// Mitsubishi GX Works2 project: ZhaoQing_FenRong_Debug   PLC: Q06UDEH

TYPE ShuttleCarIO : STRUCT
  xReady : BOOL;  (* 准备就绪 *)
  xForward : BOOL;  (* 正转 *)
  xBackward : BOOL;  (* 反转 *)
  iCurrentPos : INT;  (* 当前位置 *)
  iDestinationPos : INT;  (* 目标位置 *)
  xCW : BOOL;  (* 正转输出 *)
  xCCW : BOOL;  (* 反转输出 *)
  xBrake : BOOL;  (* 刹车 *)
  xHomeSwitch : BOOL;  (* 零位接近开关 *)
  xPosLimit : BOOL;  (* 正限位 *)
  xNegLimit : BOOL;  (* 负限位 *)
  xMDIExe : BOOL;  (* MDI开始 *)
  xMDIDone : BOOL;  (* MDI 完成 *)
  xPassLimit : BOOL;  (* 限位屏蔽 *)
  xPosLimitCatch : BOOL;  (* 正限位捕捉 *)
  xNegLimitCatch : BOOL;  (* 负限位捕捉 *)
  xHomeExe : BOOL;  (* 开始寻零 *)
  xHomeDone : BOOL;  (* 寻零完成 *)
  xHomeBusy : BOOL;  (* 寻零中 *)
  xHomeFailed : BOOL;  (* 寻零失败 *)
  xBusy : BOOL;  (* 工作中 *)
  tArriveDelay : TIME;  (* 到位延时 *)
  xCylinder : BOOL;  (* 气缸控制 *)
  tBrakeDelay : TIME;  (* 抱闸延时 *)
  xPauseRamp : BOOL;  (* 暂停减速斜坡标志位 *)
  xPresentDetect1 : BOOL;  (* 物料有无检测1 *)
  xPresentDetect2 : BOOL;  (* 物料有无检测2 *)
  xOvertimeAlarm : BOOL;  (* 超时报警 *)
  tSetOverTime : TIME;  (* 设置超时时间 *)
  xLooseDetect : BOOL;  (* 松绳检测 *)
  xLooseAlarm : BOOL;  (* 松绳报警 *)
END_STRUCT END_TYPE

TYPE SwitchIO : STRUCT
  xLiftCylinderRetractDetect : BOOL;
  xLiftCylinderExtendDetect : BOOL;
  xLiftCylinderRetract : BOOL;
  xLiftCylinderExtend : BOOL;
  xEntryBarCylinderRetract : BOOL;
  xLiftCylinderExtendInit : BOOL;
  xEntryEnable : BOOL;
  xExitEnable : BOOL;
  xExitBarCylinderRetract : BOOL;
  xSwithEnable : BOOL;
  xLiftCylinderRetractButton : BOOL;
  xLiftCylinderExtendButton : BOOL;
  xEntryBarCylinderRetractButton : BOOL;
  xExitBarCylinderRetractButton : BOOL;
END_STRUCT END_TYPE

TYPE BarCylinderIO : STRUCT
  xPresentSwitch : BOOL;  (* 行程开关 *)
  xBarCylinder : BOOL;  (* 阻挡气缸 *)
  xEmpty : BOOL;  (* 为空指示 *)
  xTransportMotorCW : BOOL;  (* 输送电机正转 *)
  xUnload : BOOL;  (* 下料 *)
  xBarCylinderButton : BOOL;  (* 阻挡气缸 *)
  xTransportMotorCWButton : BOOL;  (* 输送电机正转按钮 *)
  xLoad : BOOL;  (* 上料 *)
  xNextRun : BOOL;  (* 下位设备开始运行 *)
  xTransportMotorCCWButton : BOOL;  (* 输送电机反转按钮 *)
  xTransportMotorCCW : BOOL;  (* 输送电机反转 *)
  iProductCategory : INT;  (* 产品种类 *)
  tLoadDelay : TIME;  (* 上料延时 *)
END_STRUCT END_TYPE

TYPE ConveyorIO : STRUCT
  iProductCategory : INT;  (* 产品类型0：无料1：正极  2：负极 3：隔膜 4：空料架 *)
  xCWPresent : BOOL;  (* 正转检测有无传感器 *)
  xCCWPresent : BOOL;  (* 反转检测有无传感器 *)
  xLoad : BOOL;  (* 上料请求 *)
  xUnload : BOOL;  (* 下料请求 *)
  xMotorCW : BOOL;  (* 电机正转 *)
  xMotorCCW : BOOL;  (* 电机反转 *)
  xEmpty : BOOL;  (* 线体状态为空 *)
  xNextRun : BOOL;  (* 下段线体运行 *)
  xUnloadCCW : BOOL;  (* 下料为反转 *)
  xloadCCW : BOOL;  (* 上料为反转 *)
  xLeave : BOOL;  (* 已经离开 *)
  xForward : BOOL;  (* 正转手动 *)
  xBackward : BOOL;  (* 反转手动 *)
  xBusy : BOOL;  (* 工作中 *)
  tLoadDelay : TIME;  (* 进入延时设置 *)
  xPutInto : BOOL;  (* 线体直接投入物料 *)
  xUnloadAlarm : BOOL;  (* 下料报警 *)
  xPosLimit : BOOL;  (* 正限位 *)
  xNegLimit : BOOL;  (* 负限位 *)
  xOverWidthAlarm : BOOL;  (* 超宽报警 *)
  xLimitAlarrm : BOOL;  (* 限位报警 *)
  iDeviceID : INT;  (* 线体ID *)
  xSizeDeficientDetect : BOOL;  (* 尺寸不足检测标志位 *)
END_STRUCT END_TYPE

TYPE RGVCommunication : STRUCT
  xFullLoadRequest : BOOL;  (* 满框上料请求 *)
  xFullUnloadRequest : BOOL;  (* 满框下料请求 *)
  xEmptyLoadRequest : BOOL;  (* 空框上料请求 *)
  xEmptyUnloadRequest : BOOL;  (* 空框下料请求 *)
  xFullLoadRequestAkn : BOOL;  (* 满框上料请求确认 *)
  xFullUnloadRequestAkn : BOOL;  (* 满框下料请求确认 *)
  xEmptyLoadRequestAkn : BOOL;  (* 空框上料请求确认 *)
  xEmptyUnloadRequestAkn : BOOL;  (* 空框下料请求确认 *)
  xFullLoadComplete : BOOL;  (* 满框上料完成 *)
  xFullUnloadComplete : BOOL;  (* 满框下料完成 *)
  xEmptyLoadComplete : BOOL;  (* 空框上料完成 *)
  xEmptyUnloadComplete : BOOL;  (* 空框下料完成 *)
  xFullLoadCompleteAkn : BOOL;  (* 满框上料完成确认 *)
  xFullUnloadCompleteAkn : BOOL;  (* 满框下料完成确认 *)
  xEmptyLoadCompleteAkn : BOOL;  (* 空框上料完成确认 *)
  xEmptyUnloadCompleteAkn : BOOL;  (* 空框下料完成确认 *)
  xMdiExe : BOOL;  (* RGV 执行 *)
  xMdiDone : BOOL;  (* RGV 执行完成 *)
  iCurrentPostion : INT;  (* RGV当前位置 *)
  iDestinationPos : INT;  (* RGV目标位置 *)
  xEmpty1 : BOOL;
  xNextRun1 : BOOL;
  xEmpty2 : BOOL;
  xNextRun2 : BOOL;
  xLoad1 : BOOL;
  xUnload1 : BOOL;
  xLoad2 : BOOL;
  xUnload2 : BOOL;
  xCollisionAlarm : BOOL;  (* 干涉报警 *)
  xRemoteReset : BOOL;  (* 远程复位 *)
  xAuto : BOOL;  (* 自动 *)
END_STRUCT END_TYPE

TYPE Stub : STRUCT
  xLoadRequest : BOOL;
  xLoadRequestAkn : BOOL;
  xUnloadRequest : BOOL;
  xUnloadRequestAkn : BOOL;
END_STRUCT END_TYPE

// global labels: Global1
VAR_GLOBAL
  g_xAuto AT M11 : BOOL;
  g_xManual : BOOL;
  g_xEStop AT X33 : BOOL;
  g_xReset AT X30 : BOOL;
  g_xStackLampRed AT Y230 : BOOL;
  g_xStackLampAmber AT Y231 : BOOL;
  g_xStackLampGreen AT Y232 : BOOL;
  g_xBuzzer AT Y233 : BOOL;
  g_xStop AT M2 : BOOL;
  g_xLocalAutoStart AT M1 : BOOL;
  g_xRemoteAutoStart AT M0 : BOOL;
  g_xRemoteAuto AT M10 : BOOL;
  g_iState AT D40 : INT;
  g_iLocalAutoStep : INT;
  g_xImport1Force AT M141 : BOOL;  (* 常温库1巷道单框强制入库 *)
  g_xImport2Force AT M142 : BOOL;  (* 常温库2巷道单框强制入库 *)
  g_xImport3Force AT M143 : BOOL;  (* 常温库3巷道单框强制入库 *)
  g_xForbidLifter7 AT M146 : BOOL;  (* 禁用提升机7 *)
  g_xResetSingle AT M4 : BOOL;  (* 单线体复位 *)
  g_iDeviceIDSelect AT D0 : INT;
  g_xPause AT M3 : BOOL;  (* 暂停 *)
  g_xAlarm : BOOL;  (* 报警 *)
  g_xCommissioning : BOOL;  (* 调试模式 *)
END_VAR

// global labels: Global
VAR_GLOBAL
  g_xQuarPackageRGVComFailed : BOOL;
  g_xPassQualityDetectStation1 AT M193 : BOOL;
  g_xPassQualityDetectStation2 AT M194 : BOOL;
  g_xPassQualityDetectStation3 AT M195 : BOOL;
END_VAR

// task Task_01 (event TRUE, interval 0, priority 31): POU, Start, TCP

PROGRAM POU
VAR
  Lifter6 : ShuttleCar;
  Lifter6IO : ShuttleCarIO;
  Conveyor6 : Conveyor;
  COnveyor6IO : ConveyorIO;
  Lifter7 : ShuttleCar;
  Lifter7IO : ShuttleCarIO;
  Conveyor7 : Conveyor;
  COnveyor7IO : ConveyorIO;
  H850Conveyor9IO : ConveyorIO;
  H850Conveyor1IOTrans : ConveyorIO;
  H850Conveyor2Trans : Conveyor;
  H850Conveyor2IOTrans : ConveyorIO;
  H850Conveyor3Trans : Conveyor;
  H850Conveyor3IOTrans : ConveyorIO;
  H850Conveyor4Trans : Conveyor;
  H850Conveyor4IOTrans : ConveyorIO;
  H850Conveyor6Trans : Conveyor;
  H850Conveyor6IOTrans : ConveyorIO;
  H850Conveyor7Trans : Conveyor;
  H850Conveyor7IOTrans : ConveyorIO;
  H850Conveyor8Trans : Conveyor;
  H850Conveyor8IOTrans : ConveyorIO;
  H2500Conveyor1 : Conveyor;
  H2500Conveyor1IO : ConveyorIO;
  H850Switch1 : Switch;
  H850Switch1IO : SwitchIO;
  H850Switch1ConveyorIn : ConveyorIO;
  H850Switch1ConveyorOut : ConveyorIO;
  H850Switch2 : Switch;
  H850Switch2IO : SwitchIO;
  H850Switch2ConveyorIn : ConveyorIO;
  H850Switch2ConveyorOut : ConveyorIO;
  H850Switch3 : Switch;
  H850Switch3IO : SwitchIO;
  H850Switch3ConveyorIn : ConveyorIO;
  H850Switch3ConveyorOut : ConveyorIO;
  H850Switch4 : Switch;
  H850Switch4IO : SwitchIO;
  H850Switch4ConveyorIn : ConveyorIO;
  H850Switch4ConveyorOut : ConveyorIO;
  H850Switch5 : Switch;
  H850Switch5IO : SwitchIO;
  H850Switch5ConveyorIn : ConveyorIO;
  H850Switch5ConveyorOut : ConveyorIO;
  H850Conveyor1 : Conveyor;
  H850Conveyor1IO : ConveyorIO;
  H2500Switch : Switch;
  H2500SwitchIO : SwitchIO;
  H2500SwitchConveyorIn : ConveyorIO;
  H2500SwitchConveyorOut : ConveyorIO;
  H2500Rotor : ShuttleCar;
  H2500RotorIO : ShuttleCarIO;
  H2500RotorConveyor : Conveyor;
  H2500RotorConveyorIO : ConveyorIO;
  H850Conveyor5Trans : Conveyor;
  H850Conveyor5IOTrans : ConveyorIO;
  H850Conveyor12 : Conveyor;
  H850Conveyor12IO : ConveyorIO;
  H850Conveyor13 : Conveyor;
  H850Conveyor13IO : ConveyorIO;
  H850Rotor : ShuttleCar;
  H850RotorIO : ShuttleCarIO;
  H850RotorConveyor : Conveyor;
  H850RotorConveyorIO : ConveyorIO;
  H750Rotor : ShuttleCar;
  H750RotorIO : ShuttleCarIO;
  H750RotorConveyor : Conveyor;
  H750RotorConveyorIO : ConveyorIO;
  H850Conveyor9 : Conveyor;
  H850Conveyor1Trans : Conveyor;
  H750Switch : Switch;
  H750SwitchIO : SwitchIO;
  H750SwitchConveyorIn : ConveyorIO;
  H750SwitchConveyorOut : ConveyorIO;
  Lifter6Velocity : ShuttleCarVelocityFB;
  Lifter7Velocity : ShuttleCarVelocityFB;
  H750Conveyor1 : Conveyor;
  H750Conveyor1IO : ConveyorIO;
  H750Conveyor2 : Conveyor;
  H750Conveyor2IO : ConveyorIO;
  H750Conveyor3 : Conveyor;
  H750Conveyor3IO : ConveyorIO;
  H750Conveyor4 : Conveyor;
  H750Conveyor4IO : ConveyorIO;
  H750Conveyor5 : Conveyor;
  H750Conveyor5IO : ConveyorIO;
  H750Conveyor6 : Conveyor;
  H750Conveyor6IO : ConveyorIO;
  H750Switch1 : Switch;
  H750Switch1IO : SwitchIO;
  H750Switch1ConveyorIn : ConveyorIO;
  H750Switch1ConveyorOut : ConveyorIO;
  H750Switch2 : Switch;
  H750Switch2IO : SwitchIO;
  H750Switch2ConveyorIn : ConveyorIO;
  H750Switch2ConveyorOut : ConveyorIO;
  H750Switch3 : Switch;
  H750Switch3IO : SwitchIO;
  H750Switch3ConveyorIn : ConveyorIO;
  H750Switch3ConveyorOut : ConveyorIO;
  H2500BarCylinder : BarCylinder;
  H2500BarCylinderIO : BarCylinderIO;
  H2500EmptyASwitch : Switch;
  H2500EmptyASwitchIO : SwitchIO;
  H2500EmptyASwitchConveyorIn : ConveyorIO;
  H2500EmptyASwitchConveyorOut : ConveyorIO;
  H2500EmptyBSwitch : Switch;
  H2500EmptyBSwitchIO : SwitchIO;
  H2500EmptyBSwitchConveyorIn : ConveyorIO;
  H2500EmptyBSwitchConveyorOut : ConveyorIO;
  m_iH750Switch1Select : INT;  (* 选择入料位 *)
  H750ImportConveyor1 : Conveyor;  (* 选择入料位 *)
  H750ImportConveyor1IO : ConveyorIO;  (* 选择入料位 *)
  m_iH750Switch2Select : INT;  (* 选择入料位 *)
  m_iH750Switch3Select : INT;  (* 选择入料位 *)
  H750ImportConveyor2 : Conveyor;  (* 选择入料位 *)
  H750ImportConveyor2IO : ConveyorIO;  (* 选择入料位 *)
  H750ImportConveyor3 : Conveyor;  (* 选择入料位 *)
  H750ImportConveyor3IO : ConveyorIO;  (* 选择入料位 *)
  H750ImportConveyor4 : Conveyor;  (* 选择入料位 *)
  H750ImportConveyor4IO : ConveyorIO;  (* 选择入料位 *)
  H750ImportConveyor5 : Conveyor;  (* 选择入料位 *)
  H750ImportConveyor5IO : ConveyorIO;  (* 选择入料位 *)
  H750ImportConveyor6 : Conveyor;  (* 选择入料位 *)
  H750ImportConveyor6IO : ConveyorIO;  (* 选择入料位 *)
  H750ImportCylinder1 : ShuttleCar;
  H750ImportCylinder1IO : ShuttleCarIO;
  H750ImportCylinder2 : ShuttleCar;
  H750ImportCylinder2IO : ShuttleCarIO;
  H750ImportCylinder3 : ShuttleCar;
  H750ImportCylinder3IO : ShuttleCarIO;
  m_tonSwitch1SeleteDelay : TON;
  m_xSwitch1SeleteDelay : BOOL;
  m_tSwitch1SeleteDelayCurrentTime : TIME;
  m_tonSwitch1NOSeleteDelay : TON;
  m_xSwitch1NoSeleteDelay : BOOL;
  m_tSwitch1NOSeleteDelayCurrentTi : TIME;
  m_xH750RotorDirection : BOOL;  (* 分容出库转台旋转方向 *)
  m_tonSwitch2NOSeleteDelay : TON;
  m_xSwitch2NoSeleteDelay : BOOL;
  m_tSwitch2NOSeleteDelayCurrentTi : TIME;
  m_xSwitch2SeleteDelay : BOOL;
  m_tonSwitch3NOSeleteDelay : TON;
  m_xSwitch3NoSeleteDelay : BOOL;
  m_tSwitch3NOSeleteDelayCurrentTi : TIME;
  m_xSwitch3SeleteDelay : BOOL;
  H2500Export1Cylinder : ShuttleCar;
  H2500Export1CylinderIO : ShuttleCarIO;
  H2500Export2Cylinder : ShuttleCar;
  H2500Export2CylinderIO : ShuttleCarIO;
  H2500Export3Cylinder : ShuttleCar;
  H2500Export3CylinderIO : ShuttleCarIO;
  H2500Export1Conveyor1 : Conveyor;
  H2500Export1Conveyor1IO : ConveyorIO;
  H2500Export1Conveyor2 : Conveyor;
  H2500Export1Conveyor2IO : ConveyorIO;
  H2500Export2Conveyor1 : Conveyor;
  H2500Export2Conveyor1IO : ConveyorIO;
  H2500Export2Conveyor2 : Conveyor;
  H2500Export2Conveyor2IO : ConveyorIO;
  H2500Export3Conveyor1 : Conveyor;
  H2500Export3Conveyor1IO : ConveyorIO;
  H2500Export3Conveyor2 : Conveyor;
  H2500Export3Conveyor2IO : ConveyorIO;
  H2500Export1Switch : Switch;
  H2500Export1SwitchIO : SwitchIO;
  H2500Export1SwitchConveyorIn : ConveyorIO;
  H2500Export1SwitchConveyorOut : ConveyorIO;
  H2500Export2Switch : Switch;
  H2500Export2SwitchIO : SwitchIO;
  H2500Export2SwitchConveyorIn : ConveyorIO;
  H2500Export2SwitchConveyorOut : ConveyorIO;
  H2500Export3Switch : Switch;
  H2500Export3SwitchIO : SwitchIO;
  H2500Export3SwitchConveyorIn : ConveyorIO;
  H2500Export3SwitchConveyorOut : ConveyorIO;
  H2500Export1Conveyor3 : Conveyor;
  H2500Export1Conveyor3IO : ConveyorIO;
  H2500Export1Conveyor4 : Conveyor;
  H2500Export1Conveyor4IO : ConveyorIO;
  H2500Export2Conveyor3 : Conveyor;
  H2500Export2Conveyor3IO : ConveyorIO;
  H2500Export2Conveyor4 : Conveyor;
  H2500Export2Conveyor4IO : ConveyorIO;
  H2500Export3Conveyor3 : Conveyor;
  H2500Export3Conveyor3IO : ConveyorIO;
  H2500Export3Conveyor4 : Conveyor;
  H2500Export3Conveyor4IO : ConveyorIO;
  m_tpH2500RotorReset : TP;
  m_tH2500RotorResetCurrentTime : TIME;
  QuarPackageRGV : RGVCommunication;
  QuarPackage1Stub : Stub;
  QuarPackage2Stub : Stub;
  QuarPackage3Stub : Stub;
  QuarPackage4Stub : Stub;
  m_xDefectDetect1Complete : BOOL;
  H850Conveyor14 : Conveyor;
  H850Conveyor14IO : ConveyorIO;
  H850Switch4Task : PiorityFb;
  m_iH850Switch4Task : INT;
  m_xManualLoad : BOOL;
  m_xDefectDetect2Complete : BOOL;
  m_xDefectDetect3Complete : BOOL;
END_VAR
H850Switch1(ConveyorEntryIO:=H850Switch1ConveyorIn ,
                                                        ConveyorExitIO:=H850Switch1ConveyorOut ,
                                                        SwitchIO:=H850Switch1IO );
H850Switch1IO.xLiftCylinderExtendButton:=M30;
H850Switch1IO.xLiftCylinderRetractButton:=M31;
H850Switch1IO.xExitBarCylinderRetractButton:=M32;
Y260:=H850Switch1IO.xEXITBarCylinderRetract;
Y25E:=H850Switch1IO.xLiftCylinderExtend;
Y25D:=H850Switch1IO.xLiftCylinderRetract;
H850Switch1IO.xLiftCylinderExtendDetect:=X5D;
H850Switch1IO.xLiftCylinderRetractDetect:=X5E;
H850Switch1ConveyorIn.xForward:=M33;
H850Switch1ConveyorIn.xCWPresent:=X60;
H850Switch1ConveyorIn.iDeviceID:=12110;
Y269:=H850Switch1ConveyorIn.xMotorCW OR H850Switch2ConveyorIn.xMotorCW;
H850Switch1ConveyorOut.xForward:=M34;
H850Switch1ConveyorOut.xCWPresent:=X5F;
Y25F:=H850Switch1ConveyorOut.xMotorCW;
H850Switch1ConveyorOut.iDeviceID:=12110;

H850Switch2(ConveyorEntryIO:=H850Switch2ConveyorIn ,
                                                        ConveyorExitIO:=H850Switch2ConveyorOut ,
                                                        SwitchIO:=H850Switch2IO );
H850Switch2IO.xLiftCylinderExtendButton:=M35;
H850Switch2IO.xLiftCylinderRetractButton:=M36;
H850Switch2IO.xExitBarCylinderRetractButton:=M37;
Y128:=H850Switch2IO.xEXITBarCylinderRetract;
Y262:=H850Switch2IO.xLiftCylinderExtend;
Y261:=H850Switch2IO.xLiftCylinderRetract;
H850Switch2IO.xLiftCylinderExtendDetect:=X61;
H850Switch2IO.xLiftCylinderRetractDetect:=X62;
H850Switch2ConveyorIn.xForward:=M38;
H850Switch2ConveyorIn.tLoadDelay:=T#2s500ms;
H850Switch2ConveyorIn.xCWPresent:=X63;
H850Switch2ConveyorIn.iDeviceID:=12110;
(*Y187:=H850Switch2ConveyorIn.xMotorCW;*)
H850Switch2ConveyorOut.xForward:=M39;
H850Switch2ConveyorOut.xCWPresent:=X6A;
Y263:=H850Switch2ConveyorOut.xMotorCW;
H850Switch2ConveyorOut.iDeviceID:=12110;

H850Switch3(ConveyorEntryIO:=H850Switch3ConveyorIn ,
                                                        ConveyorExitIO:=H850Switch3ConveyorOut ,
                                                        SwitchIO:=H850Switch3IO );
H850Switch3IO.xLiftCylinderExtendButton:=M40;
H850Switch3IO.xLiftCylinderRetractButton:=M41;
H850Switch3IO.xExitBarCylinderRetractButton:=M42;
Y128:=H850Switch3IO.xEXITBarCylinderRetract;
Y265:=H850Switch3IO.xLiftCylinderExtend;
Y266:=H850Switch3IO.xLiftCylinderRetract;
H850Switch3IO.xLiftCylinderExtendDetect:=X66;
H850Switch3IO.xLiftCylinderRetractDetect:=X65;
H850Switch3ConveyorIn.xForward:=M43;
H850Switch3ConveyorIn.xCWPresent:=X68;
H850Switch3ConveyorIn.tLoadDelay:=T#1s;
Y267:=H850Switch3ConveyorIn.xMotorCW;
H850Switch3ConveyorIn.iDeviceID:=12109;
H850Switch3ConveyorOut.xForward:=M44;
H850Switch3ConveyorOut.xCWPresent:=X67;
Y268:=H850Switch3ConveyorOut.xMotorCW;
H850Switch3IO.xLiftCylinderExtendInit:=1;
H850Switch3ConveyorOut.iDeviceID:=12109;

H850Switch4(ConveyorEntryIO:=h850Conveyor12IO,
                                                        ConveyorExitIO:=H850Switch4ConveyorOut ,
                                                        SwitchIO:=H850Switch4IO );
H850Switch4IO.xLiftCylinderExtendButton:=M45;
H850Switch4IO.xLiftCylinderRetractButton:=M46;
H850Switch4IO.xExitBarCylinderRetractButton:=M47;
Y128:=H850Switch4IO.xEXITBarCylinderRetract;
Y272:=H850Switch4IO.xLiftCylinderExtend;
Y270:=H850Switch4IO.xLiftCylinderRetract;
H850Switch4IO.xLiftCylinderExtendDetect:=X6F;
H850Switch4IO.xLiftCylinderRetractDetect:=X70;
H850Switch4ConveyorIn.xForward:=M48;
H850Switch4ConveyorIn.xCWPresent:=X131;
H850Switch4ConveyorIn.iDeviceID:=12301;
(*Y187:=H850Switch4ConveyorIn.xMotorCW;*)
H850Switch4ConveyorOut.xForward:=M49;
H850Switch4ConveyorOut.xCWPresent:=X131;
Y30B:=H850Switch4ConveyorOut.xMotorCW ;
H850Switch4ConveyorOut.iDeviceID:=12301;

H850Switch5(ConveyorEntryIO:=H850Switch5ConveyorIn ,
                                                        ConveyorExitIO:=H850Switch5ConveyorOut ,
                                                        SwitchIO:=H850Switch5IO );
H850Switch5IO.xLiftCylinderExtendButton:=M50;
H850Switch5IO.xLiftCylinderRetractButton:=M51;
H850Switch5IO.xExitBarCylinderRetractButton:=M52;
Y128:=H850Switch5IO.xEXITBarCylinderRetract;
Y274:=H850Switch5IO.xLiftCylinderExtend;
Y271:=H850Switch5IO.xLiftCylinderRetract;
H850Switch5IO.xLiftCylinderExtendDetect:=X71;
H850Switch5IO.xLiftCylinderRetractDetect:=X72;
H850Switch5ConveyorIn.xForward:=M53;
H850Switch5ConveyorIn.xCWPresent:=X130;
Y30A:=H850Switch5ConveyorIn.xMotorCW;
H850Switch5ConveyorIn.iDeviceID:=12302;
H850Switch5ConveyorOut.xForward:=M54;
H850Switch5ConveyorOut.xCWPresent:=X130;
Y26C:=H850Switch5ConveyorOut.xMotorCW AND NOT Y26F;(*同一电机互锁反转信号*)
H850Switch5ConveyorOut.iDeviceID:=12302;

Lifter6(ShuttleCarInOut:=Lifter6IO);
ShuttleCarCurrentPosition( X3C OR X3D ,X3C ,X3D, FALSE, Lifter6IO.iCurrentPos );
Lifter6Velocity(xEnable:= g_xAuto ,
                          xMotorCW:= Lifter6IO.xCW ,
                          xMotorCCW:= Lifter6IO.xCCW,
                          xPosition1Switch:= X3C ,
                          xDecelerationSwitch:= X5B ,
	                      xPosition2Switch:= X3D ,
	                      xHighSpeed:= Y23E );
Lifter6IO.xReady:=X2C;
Lifter6Io.xForward:=M55 OR X41;
Lifter6IO.xBackward:=M56 OR X42;
Lifter6IO.xPosLimit:=X3E;
Lifter6IO.xNegLimit:=X3F;
Lifter6IO.xLooseDetect:=X40;
M177:=Lifter6IO.xLooseAlarm;
Y23D:=Lifter6IO.xCW;
Y23C:=Lifter6IO.xCCW;
Y241:=Lifter6IO.xBrake;

Conveyor6(ConveyorMotor:=Conveyor6IO);
Conveyor6IO.xForward:=M57;
Conveyor6IO.xBackward:=M58;
Conveyor6IO.xCWPresent:=X43;
Conveyor6IO.xCCWPresent:=X44;
Y24B:=Conveyor6IO.xMotorCW;
Y24C:=Conveyor6IO.xMotorCCW;
COnveyor6IO.xloadCCW:=1;
COnveyor6IO.iDeviceID:=6;

Lifter7(ShuttleCarInOut:=Lifter7IO);
ShuttleCarCurrentPosition( X45 OR X46 ,X45 ,X46, FALSE, Lifter7IO.iCurrentPos );
Lifter7Velocity(xEnable:= g_xAuto ,
                          xMotorCW:= Lifter7IO.xCW ,
                          xMotorCCW:= Lifter7IO.xCCW,
                          xPosition1Switch:= X45 ,
                          xDecelerationSwitch:= X5C ,
	                      xPosition2Switch:= X46 ,
	                      xHighSpeed:= Y244 );
Lifter7IO.xReady:=X2D;
Lifter7Io.xForward:=M59 OR X4A;
Lifter7IO.xBackward:=M60 OR X4B;
Lifter7IO.xLooseDetect:=X49;
M178:=Lifter7IO.xLooseAlarm;
Lifter7IO.xPosLimit:=X47;
Lifter7IO.xNegLimit:=X48;
Y243:=Lifter7IO.xCW;
Y242:=Lifter7IO.xCCW;
Y247:=Lifter7IO.xBrake;

Conveyor7(ConveyorMotor:=Conveyor7IO);
Conveyor7IO.xForward:=M61;
Conveyor7IO.xBackward:=M62;
Conveyor7IO.xCWPresent:=X4D;
Conveyor7IO.xCCWPresent:=X4C;
Y24D:=Conveyor7IO.xMotorCW;
(*:=Conveyor7IO.xMotorCCW;*)
Conveyor7IO.xSizeDeficientDetect:=1; (*尺寸检测*)
M184:=Conveyor7IO.xOverWidthAlarm;
Conveyor7IO.tLoadDelay:=T#500ms;
COnveyor7IO.iDeviceID:=7;

H850Conveyor1(ConveyorMotor:=H850Conveyor1IO);
(*H850Conveyor1IO.tLeaveDelay:=t#2s;*)
H850Conveyor1IO.xForward:=M63;
H850Conveyor1IO.xCWPresent:=X73;
Y273:=H850Conveyor1IO.xMotorCW;
H850Conveyor1IO.iDeviceID:=12114;

H850Conveyor12(ConveyorMotor:=H850Conveyor12IO);
H850Conveyor12IO.xForward:=M82;
H850Conveyor12IO.xCWPresent:=X131(*X6D*);
Y26D:=H850Conveyor12IO.xMotorCW;
H850Conveyor12IO.iDeviceID:=12111;

H850Conveyor13(ConveyorMotor:=H850Conveyor13IO);
H850Conveyor13IO.xForward:=M83;
H850Conveyor13IO.xCWPresent:=X6E;
Y26E:=H850Conveyor13IO.xMotorCW;
H850Conveyor13IO.iDeviceID:=12112;

H850Conveyor14(ConveyorMotor:=H850Conveyor14IO);
H850Conveyor14IO.xForward:=M192;
H850Conveyor14IO.xCWPresent:=X13B;
Y26F:=H850Conveyor14IO.xMotorCCW AND NOT Y26C;(*同一个电机互锁正转信号*)
H850Conveyor14IO.iDeviceID:=12113;
H850Conveyor14IO.xUnloadCCW:=1;
H850Conveyor14Io.tLoadDelay:=T#2s;

H2500Conveyor1(ConveyorMotor:=H2500Conveyor1IO);
H2500Conveyor1IO.xForward:=M64;
H2500Conveyor1IO.xCWPresent:=X7D;
Y27D:=H2500Conveyor1IO.xMotorCW;
H2500Conveyor1IO.iDeviceID:=12116;

H2500Switch(ConveyorEntryIO:=H2500SwitchConveyorIn ,
                                                        ConveyorExitIO:=H2500SwitchConveyorOut ,
                                                        SwitchIO:=H2500SwitchIO );
H2500SwitchIO.xLiftCylinderExtendButton:=M65;
H2500SwitchIO.xLiftCylinderRetractButton:=M66;
H2500SwitchIO.xExitBarCylinderRetractButton:=M67;
Y128:=H2500SwitchIO.xEXITBarCylinderRetract;
Y27E:=H2500SwitchIO.xLiftCylinderExtend;
Y27F:=H2500SwitchIO.xLiftCylinderRetract;
H2500SwitchIO.xLiftCylinderExtendDetect:=X7E;
H2500SwitchIO.xLiftCylinderRetractDetect:=X7F;
H2500SwitchConveyorIn.xForward:=M68;
H2500SwitchConveyorIn.xCWPresent:=X80;
H2500SwitchConveyorIn.tLoadDelay:=T#2s;
Y280:=H2500SwitchConveyorIn.xMotorCW;
H2500SwitchConveyorIn.iDeviceID:=12204;
H2500SwitchConveyorOut.xForward:=M84;
H2500SwitchConveyorOut.xCWPresent:=X80;
Y281:=H2500SwitchConveyorOut.xMotorCW OR H2500BarCylinderIO.xTransportMotorCW  ;(*倍速链线体*)
Y2F3:=H2500SwitchConveyorOut.xMotorCW OR H2500BarCylinderIO.xTransportMotorCW ;(*滚筒线1*)
Y2F4:=H2500SwitchConveyorOut.xMotorCW OR H2500BarCylinderIO.xTransportMotorCW ;(*滚筒线2*)
H2500SwitchConveyorOut.iDeviceID:=12204;

H2500BarCylinder(BarCylinderIO:=H2500BarCylinderIO);
H2500BarCylinderIO.xBarCylinderButton:=M196;
H2500BarCylinderIO.xPresentSwitch:=X82;
Y283:=H2500BarCylinderIO.xBarCylinder;

H2500Rotor(ShuttleCarInOut:=H2500RotorIO);
ShuttleCarCurrentPosition( X83 OR X84 ,X83 ,X84, FALSE,H2500RotorIO.iCurrentPos );
H2500RotorIO.xReady:=X2E;
H2500RotorIO.xForward:=M70 ;
H2500RotorIO.xBackward:=M71 ;
H2500RotorIO.xPosLimit:=X85;
H2500RotorIO.xNegLimit:=X86;
Y284:=H2500RotorIO.xCW;
Y285:=H2500RotorIO.xCCW;
Y295:=H2500RotorIO.xBrake;

H2500RotorConveyor(ConveyorMotor:=H2500RotorConveyorIO);
H2500RotorConveyorIO.xForward:=M72;
H2500RotorConveyorIO.xBackward:=M73;
H2500RotorConveyorIO.xCWPresent:=X88;
H2500RotorConveyorIO.xCCWPresent:=X87;
Y286:=H2500RotorConveyorIO.xMotorCW;
Y287:=H2500RotorConveyorIO.xMotorCCW;
H2500RotorConveyorIO.tLoadDelay:=T#1s500ms;
H2500RotorConveyorIO.iDeviceID:=12502;

H850Conveyor1Trans(ConveyorMotor:=H850Conveyor1IOTrans);
H850Conveyor1IOTrans.xForward:=M74;
H850Conveyor1IOTrans.xCWPresent:=X75;
Y275:=H850Conveyor1IOTrans.xMotorCW;
H850Conveyor1IOTrans.iDeviceID:=12101;

H850Conveyor2Trans(ConveyorMotor:=H850Conveyor2IOTrans);
H850Conveyor2IOTrans.xForward:=M75;
H850Conveyor2IOTrans.xCWPresent:=X76;
Y276:=H850Conveyor2IOTrans.xMotorCW;
H850Conveyor2IOTrans.iDeviceID:=12102;

H850Conveyor3Trans(ConveyorMotor:=H850Conveyor3IOTrans);
H850Conveyor3IOTrans.xForward:=M76;
H850Conveyor3IOTrans.xCWPresent:=  X77;
Y277:=H850Conveyor3IOTrans.xMotorCW;
H850Conveyor3IOTrans.iDeviceID:=12103;

H850Conveyor4Trans(ConveyorMotor:=H850Conveyor4IOTrans);
H850Conveyor4IOTrans.xForward:=M77;
H850Conveyor4IOTrans.xCWPresent:=X78;
Y278:=H850Conveyor4IOTrans.xMotorCW;
H850Conveyor4IOTrans.iDeviceID:=12104;

H850Conveyor5Trans(ConveyorMotor:=H850Conveyor5IOTrans);
H850Conveyor5IOTrans.xForward:=M78;
H850Conveyor5IOTrans.xCWPresent:=X79;
Y279:=H850Conveyor5IOTrans.xMotorCW;
H850Conveyor5IOTrans.iDeviceID:=12105;		

H850Conveyor6Trans(ConveyorMotor:=H850Conveyor6IOTrans);
H850Conveyor6IOTrans.xForward:=M79;
H850Conveyor6IOTrans.xCWPresent:=X7A;
Y27A:=H850Conveyor6IOTrans.xMotorCW;
H850Conveyor6IOTrans.iDeviceID:=12106;

H850Conveyor7Trans(ConveyorMotor:=H850Conveyor7IOTrans);
H850Conveyor7IOTrans.xForward:=M80;
H850Conveyor7IOTrans.xCWPresent:=X7B;
Y27B:=H850Conveyor7IOTrans.xMotorCW;
H850Conveyor7IOTrans.iDeviceID:=12107;

H850Conveyor8Trans(ConveyorMotor:=H850Conveyor8IOTrans);
H850Conveyor8IOTrans.xForward:=M81;
H850Conveyor8IOTrans.xCWPresent:=X7C;
Y27C:=H850Conveyor8IOTrans.xMotorCW;
H850Conveyor8IOTrans.iDeviceID:=12108;

H850Rotor(ShuttleCarInOut:=H850RotorIO);
ShuttleCarCurrentPosition( X38 OR X39 ,X39 ,X38, FALSE, H850RotorIO.iCurrentPos );
H850RotorIO.xReady:=X2B;
H850RotorIO.xForward:=M85;
H850RotorIO.xBackward:=M86;
H850RotorIO.xPosLimit:=X37;
H850RotorIO.xNegLimit:=X36;
Y238:=H850RotorIO.xCW;
Y239:=H850RotorIO.xCCW;
Y237:=H850RotorIO.xBrake;
H850RotorIO.xPassLimit:=M29;

H850RotorConveyor(ConveyorMotor:=H850RotorConveyorIO);
H850RotorConveyorIO.xForward:=M87;
H850RotorConveyorIO.xBackward:=M105;
H850RotorConveyorIO.xCWPresent:=X3A;
H850RotorConveyorIO.xCCWPresent:=X35;
Y25B:=H850RotorConveyorIO.xMotorCW;
Y23A:=H850RotorConveyorIO.xMotorCCW;
H850RotorConveyorIO.xUnloadCCW:=1;
H850RotorConveyorIO.iDeviceID:=12501;

H850Conveyor9(ConveyorMotor:=H850Conveyor9IO);
H850Conveyor9IO.xForward:=M89;
H850Conveyor9IO.xCWPresent:=X3B;
Y23B:=H850Conveyor9IO.xMotorCW;
H850Conveyor9IO.iDeviceID:=12148;

H750Rotor(ShuttleCarInOut:=H750RotorIO);
ShuttleCarCurrentPosition( X89 OR X8A OR X135 ,X8A ,X135, X89, H750RotorIO.iCurrentPos );
H750RotorIO.xReady:=X2F;
H750RotorIO.xForward:=M90;
H750RotorIO.xBackward:=M91;
H750RotorIO.xPosLimit:=X8B;
H750RotorIO.xNegLimit:=X8C;
Y28A:=H750RotorIO.xCW;
Y289:=H750RotorIO.xCCW;
Y28E:=H750RotorIO.xBrake;
H750RotorIO.tArriveDelay:=T#200ms;

H750RotorConveyor(ConveyorMotor:=H750RotorConveyorIO);
H750RotorConveyorIO.xForward:=M92;
H750RotorConveyorIO.xBackward:=M139;
H750RotorConveyorIO.xCWPresent:=X8D;
H750RotorConveyorIO.xCCWPresent:=X8E;
Y28C:=H750RotorConveyorIO.xMotorCW;
Y28B:=H750RotorConveyorIO.xMotorCCW;
H750RotorConveyorIO.iDeviceID:=12503;

H750Switch(ConveyorEntryIO:=H750SwitchConveyorIn,
                         ConveyorExitIO:=H750SwitchConveyorOut,
                        SwitchIO:=H750SwitchIO );
H750SwitchIO.xLiftCylinderExtendButton:=M93;
H750SwitchIO.xLiftCylinderRetractButton:=M94;
Y290:=H750SwitchIO.xLiftCylinderExtend;
Y28F:=H750SwitchIO.xLiftCylinderRetract;
H750SwitchIO.xLiftCylinderExtendDetect:=X8F;
H750SwitchIO.xLiftCylinderRetractDetect:=X90;
H750SwitchConveyorIn.xForward:=M95;
H750SwitchConveyorIn.xCWPresent:=X93;
Y288:=H750SwitchConveyorIn.xMotorCW;
Y2F2:=H750SwitchConveyorIn.xMotorCW;
H750SwitchConveyorIn.iDeviceID:=12118;
H750SwitchConveyorIn.tLoadDelay:=T#2s;
H750SwitchConveyorOut.xForward:=M96;
H750SwitchConveyorOut.xCWPresent:=X91;
Y291:=H750SwitchConveyorOut.xMotorCW;
H750SwitchIO.xLiftCylinderExtendInit:=0;
H750SwitchConveyorOut.iDeviceID:=12207;

H750Conveyor1(ConveyorMotor:=H750Conveyor1IO);
H750Conveyor1IO.xForward:=M108;
H750Conveyor1IO.xCWPresent:=X98;
Y298:=H750Conveyor1IO.xMotorCW;
H750Conveyor1IO.iDeviceID:=12119;

H750Conveyor2(ConveyorMotor:=H750Conveyor2IO);
H750Conveyor2IO.xForward:=M109;
H750Conveyor2IO.xCWPresent:=X99;
Y299:=H750Conveyor2IO.xMotorCW;
H750Conveyor2IO.iDeviceID:=12120;
(********1巷道*************)
H750Switch1(ConveyorEntryIO:=H750Switch1ConveyorIn,
                         ConveyorExitIO:=H750Switch1ConveyorOut,
                        SwitchIO:=H750Switch1IO );
H750Switch1IO.xLiftCylinderExtendButton:=M114;
H750Switch1IO.xLiftCylinderRetractButton:=M115;
H750Switch1IO.xExitBarCylinderRetractButton:=M136;
Y29E:=H750Switch1IO.xLiftCylinderExtend;
Y29D:=H750Switch1IO.xLiftCylinderRetract;
Y29B:= NOT (H750Switch1IO.xExitBarCylinderRetract OR m_iH750Switch1Select=2 ) ;
Y29C:=NOT H750Switch1IO.xExitBarCylinderRetract ;
H750Switch1IO.xLiftCylinderExtendDetect:=XA4;
H750Switch1IO.xLiftCylinderRetractDetect:=XA3;
H750Switch1ConveyorIn.xForward:=M116;
H750Switch1ConveyorIn.xCWPresent:=((m_iH750Switch1Select=1 OR m_iH750Switch1Select=0)  AND  X9B) OR (m_iH750Switch1Select=2 AND X9C);
Y297:=H750Switch1ConveyorIn.xMotorCW;
H750Switch1ConveyorIn.iDeviceID:=12121;
H750Switch1ConveyorIn.tLoadDelay:=T#2s;
H750Switch1ConveyorOut.xForward:=M117;
H750Switch1ConveyorOut.xCWPresent:=((m_iH750Switch1Select=1 OR m_iH750Switch1Select=0) AND  X9B) OR (m_iH750Switch1Select=2 AND X9C);
Y2B5:=H750Switch1ConveyorOut.xMotorCW;
H750Switch1IO.xLiftCylinderExtendInit:=0;
H750Switch1ConveyorOut.iDeviceID:=12122;

H750ImportConveyor1(ConveyorMotor:=H750ImportConveyor1IO);
H750ImportConveyor1IO.xForward:=M135;
H750ImportConveyor1IO.xCWPresent:=XC3;
Y2B4:=H750ImportConveyor1IO.xMotorCW;
H750ImportConveyor1IO.tLoadDelay:=t#2S;
H750ImportConveyor1IO.iDeviceID:=12123;

H750ImportConveyor2(ConveyorMotor:=H750ImportConveyor2IO);
H750ImportConveyor2IO.xForward:=M118;
H750ImportConveyor2IO.xCWPresent:=XC5;
Y2B6:=H750ImportConveyor2IO.xMotorCW;
H750ImportConveyor2IO.tLoadDelay:=t#2S;
H750ImportConveyor2IO.iDeviceID:=12124;

H750ImportCylinder1(ShuttleCarInOut:= H750ImportCylinder1IO );
ShuttleCarCurrentPosition( XC6 OR XC7 ,XC7 ,XC6, FALSE, H750ImportCylinder1IO.iCurrentPos );
H750ImportCylinder1IO.xReady:=1;
H750ImportCylinder1IO.xForward:=M119;
H750ImportCylinder1IO.xBackward:=M120;
H750ImportCylinder1IO.xPosLimit:=1;
H750ImportCylinder1IO.xNegLimit:=1;
Y2B9:=H750ImportCylinder1IO.xCW;
Y2B8:=H750ImportCylinder1IO.xCCW;
H750ImportCylinder1IO.xCylinder:=1;

H750Conveyor3(ConveyorMotor:=H750Conveyor3IO);
H750Conveyor3IO.xForward:=M110;
H750Conveyor3IO.xCWPresent:=XA7;
Y2A2:=H750Conveyor3IO.xMotorCW;
H750Conveyor3IO.iDeviceID:=12125;

H750Conveyor4(ConveyorMotor:=H750Conveyor4IO);
H750Conveyor4IO.xForward:=M111;
H750Conveyor4IO.xCWPresent:=XA8;
Y2A3:=H750Conveyor4IO.xMotorCW;
H750Conveyor4IO.iDeviceID:=12126;
(********2巷道*************)
H750Switch2(ConveyorEntryIO:=H750Switch2ConveyorIn,
                         ConveyorExitIO:=H750Switch2ConveyorOut,
                        SwitchIO:=H750Switch2IO );
H750Switch2IO.xLiftCylinderExtendButton:=M121;
H750Switch2IO.xLiftCylinderRetractButton:=M122;
H750Switch2IO.xExitBarCylinderRetractButton:=M137;
Y2A5:=NOT (H750Switch2IO.xExitBarCylinderRetract OR m_iH750Switch2Select=2 );
Y2A6:=NOT H750Switch2IO.xExitBarCylinderRetract;
Y2A8:=H750Switch2IO.xLiftCylinderExtend;
Y2A7:=H750Switch2IO.xLiftCylinderRetract;
H750Switch2IO.xLiftCylinderExtendDetect:=XB2;
H750Switch2IO.xLiftCylinderRetractDetect:=XB3;
H750Switch2ConveyorIn.xForward:=M123;
H750Switch2ConveyorIn.xCWPresent:=((m_iH750Switch2Select=1 OR m_iH750Switch2Select=0)  AND  XAA) OR (m_iH750Switch2Select=2 AND XAB);
Y2A1:=H750Switch2ConveyorIn.xMotorCW;
H750Switch2ConveyorIn.tLoadDelay:=T#3s;
H750Switch2ConveyorIn.iDeviceID:=12127;
H750Switch2ConveyorOut.xForward:=M124;
H750Switch2ConveyorOut.xCWPresent:=((m_iH750Switch2Select=1 OR m_iH750Switch2Select=0) AND  XAA) OR (m_iH750Switch2Select=2 AND XAB);
Y2BB:=H750Switch2ConveyorOut.xMotorCW;
H750Switch2IO.xLiftCylinderExtendInit:=0;
H750Switch2ConveyorOut.iDeviceID:=12128;

H750ImportConveyor3(ConveyorMotor:=H750ImportConveyor3IO);
H750ImportConveyor3IO.xForward:=M125;
H750ImportConveyor3IO.xCWPresent:=XCA;
Y2BA:=H750ImportConveyor3IO.xMotorCW;
H750ImportConveyor3IO.tLoadDelay:=t#2S;
H750ImportConveyor3IO.iDeviceID:=12129;

H750ImportConveyor4(ConveyorMotor:=H750ImportConveyor4IO);
H750ImportConveyor4IO.xForward:=M126;
H750ImportConveyor4IO.xCWPresent:=XCC;
Y2BC:=H750ImportConveyor4IO.xMotorCW;
H750ImportConveyor4IO.tLoadDelay:=t#2S;
H750ImportConveyor4IO.iDeviceID:=12130;